// TIA Portal project "ProjektZaliczenie" (V13) (continued)
HMI tags "Default tag table"
   "Player1DataBlock_SelectedSize" : Int, 100 ms
   "Player1DataBlock_Orientation" : Bool, 100 ms
   "Player1DataBlock_ResetAll" : Bool, 100 ms
   "Player1DataBlock_Ready" : Bool, 100 ms
   "Player1DataBlock_SelectedPosition" : Int, 100 ms
   "Player1DataBlock_FieldsTypes" : Array [0..99] of Int, 100 ms
   "Player1DataBlock_Size4Count" : Int, 100 ms
   "Player1DataBlock_Size3Count" : Int, 100 ms
   "Player1DataBlock_Size2Count" : Int, 100 ms
   "Player1DataBlock_Size1Count" : Int, 100 ms
   "Player1DataBlock_ShipsReady" : Bool, 100 ms
   "Tag_ScreenNumber" : UInt, internal
   "MainDataBlock_Turn" : Bool, 100 ms
   "MainDataBlock_GameResult" : Int, 100 ms
   "Player1DataBlock_EnemyBoard{0}" : Int, 100 ms
   "Player1DataBlock_EnemyBoard{1}" : Int, 100 ms
   "Player1DataBlock_EnemyBoard{2}" : Int, 100 ms
   "Player1DataBlock_EnemyBoard{3}" : Int, 100 ms
   "Player1DataBlock_EnemyBoard{4}" : Int, 100 ms
   "Player1DataBlock_EnemyBoard{5}" : Int, 100 ms
   "Player1DataBlock_EnemyBoard{6}" : Int, 100 ms
   "Player1DataBlock_EnemyBoard{7}" : Int, 100 ms
   "Player1DataBlock_EnemyBoard{8}" : Int, 100 ms
   "Player1DataBlock_EnemyBoard{9}" : Int, 100 ms
   "Player1DataBlock_EnemyBoard{10}" : Int, 100 ms
   "Player1DataBlock_EnemyBoard{11}" : Int, 100 ms
   "Player1DataBlock_EnemyBoard{12}" : Int, 100 ms
   "Player1DataBlock_EnemyBoard{13}" : Int, 100 ms
   "Player1DataBlock_EnemyBoard{14}" : Int, 100 ms
   "Player1DataBlock_EnemyBoard{15}" : Int, 100 ms
   "Player1DataBlock_EnemyBoard{16}" : Int, 100 ms
   "Player1DataBlock_EnemyBoard{17}" : Int, 100 ms
   "Player1DataBlock_EnemyBoard{18}" : Int, 100 ms
   "Player1DataBlock_EnemyBoard{19}" : Int, 100 ms
   "Player1DataBlock_EnemyBoard{20}" : Int, 100 ms
   "Player1DataBlock_EnemyBoard{21}" : Int, 100 ms
   "Player1DataBlock_EnemyBoard{22}" : Int, 100 ms
   "Player1DataBlock_EnemyBoard{23}" : Int, 100 ms
   "Player1DataBlock_EnemyBoard{24}" : Int, 100 ms
   "Player1DataBlock_EnemyBoard{25}" : Int, 100 ms
   "Player1DataBlock_EnemyBoard{26}" : Int, 100 ms
   "Player1DataBlock_EnemyBoard{27}" : Int, 100 ms
   "Player1DataBlock_EnemyBoard{28}" : Int, 100 ms
   "Player1DataBlock_EnemyBoard{29}" : Int, 100 ms
   "Player1DataBlock_EnemyBoard{30}" : Int, 100 ms
   "Player1DataBlock_EnemyBoard{31}" : Int, 100 ms
   "Player1DataBlock_EnemyBoard{32}" : Int, 100 ms
   "Player1DataBlock_EnemyBoard{33}" : Int, 100 ms
   "Player1DataBlock_EnemyBoard{34}" : Int, 100 ms
   "Player1DataBlock_EnemyBoard{35}" : Int, 100 ms
   "Player1DataBlock_EnemyBoard{36}" : Int, 100 ms
   "Player1DataBlock_EnemyBoard{37}" : Int, 100 ms
   "Player1DataBlock_EnemyBoard{38}" : Int, 100 ms
   "Player1DataBlock_EnemyBoard{39}" : Int, 100 ms
   "Player1DataBlock_EnemyBoard{40}" : Int, 100 ms
   "Player1DataBlock_EnemyBoard{41}" : Int, 100 ms
   "Player1DataBlock_EnemyBoard{42}" : Int, 100 ms
   "Player1DataBlock_EnemyBoard{43}" : Int, 100 ms
   "Player1DataBlock_EnemyBoard{44}" : Int, 100 ms
   "Player1DataBlock_EnemyBoard{45}" : Int, 100 ms
   "Player1DataBlock_EnemyBoard{46}" : Int, 100 ms
   "Player1DataBlock_EnemyBoard{47}" : Int, 100 ms
   "Player1DataBlock_EnemyBoard{48}" : Int, 100 ms
   "Player1DataBlock_EnemyBoard{49}" : Int, 100 ms
   "Player1DataBlock_EnemyBoard{50}" : Int, 100 ms
   "Player1DataBlock_EnemyBoard{51}" : Int, 100 ms
   "Player1DataBlock_EnemyBoard{52}" : Int, 100 ms
   "Player1DataBlock_EnemyBoard{53}" : Int, 100 ms
   "Player1DataBlock_EnemyBoard{54}" : Int, 100 ms
   "Player1DataBlock_EnemyBoard{55}" : Int, 100 ms
   "Player1DataBlock_EnemyBoard{56}" : Int, 100 ms
   "Player1DataBlock_EnemyBoard{57}" : Int, 100 ms
   "Player1DataBlock_EnemyBoard{58}" : Int, 100 ms
   "Player1DataBlock_EnemyBoard{59}" : Int, 100 ms
   "Player1DataBlock_EnemyBoard{60}" : Int, 100 ms
   "Player1DataBlock_EnemyBoard{61}" : Int, 100 ms
   "Player1DataBlock_EnemyBoard{62}" : Int, 100 ms
   "Player1DataBlock_EnemyBoard{63}" : Int, 100 ms
   "Player1DataBlock_EnemyBoard{64}" : Int, 100 ms
   "Player1DataBlock_EnemyBoard{65}" : Int, 100 ms
   "Player1DataBlock_EnemyBoard{66}" : Int, 100 ms
   "Player1DataBlock_EnemyBoard{67}" : Int, 100 ms
   "Player1DataBlock_EnemyBoard{68}" : Int, 100 ms
   "Player1DataBlock_EnemyBoard{69}" : Int, 100 ms
   "Player1DataBlock_EnemyBoard{70}" : Int, 100 ms
   "Player1DataBlock_EnemyBoard{71}" : Int, 100 ms
   "Player1DataBlock_EnemyBoard{72}" : Int, 100 ms
   "Player1DataBlock_EnemyBoard{73}" : Int, 100 ms
   "Player1DataBlock_EnemyBoard{74}" : Int, 100 ms
   "Player1DataBlock_EnemyBoard{75}" : Int, 100 ms
   "Player1DataBlock_EnemyBoard{76}" : Int, 100 ms
   "Player1DataBlock_EnemyBoard{77}" : Int, 100 ms
   "Player1DataBlock_EnemyBoard{78}" : Int, 100 ms
   "Player1DataBlock_EnemyBoard{79}" : Int, 100 ms
   "Player1DataBlock_EnemyBoard{80}" : Int, 100 ms
   "Player1DataBlock_EnemyBoard{81}" : Int, 100 ms
   "Player1DataBlock_EnemyBoard{82}" : Int, 100 ms
   "Player1DataBlock_EnemyBoard{83}" : Int, 100 ms
   "Player1DataBlock_EnemyBoard{84}" : Int, 100 ms
   "Player1DataBlock_EnemyBoard{85}" : Int, 100 ms
   "Player1DataBlock_EnemyBoard{86}" : Int, 100 ms
   "Player1DataBlock_EnemyBoard{87}" : Int, 100 ms
   "Player1DataBlock_EnemyBoard{88}" : Int, 100 ms
   "Player1DataBlock_EnemyBoard{89}" : Int, 100 ms
   "Player1DataBlock_EnemyBoard{90}" : Int, 100 ms
   "Player1DataBlock_EnemyBoard{91}" : Int, 100 ms
   "Player1DataBlock_EnemyBoard{92}" : Int, 100 ms
   "Player1DataBlock_EnemyBoard{93}" : Int, 100 ms
   "Player1DataBlock_EnemyBoard{94}" : Int, 100 ms
   "Player1DataBlock_EnemyBoard{95}" : Int, 100 ms
   "Player1DataBlock_EnemyBoard{96}" : Int, 100 ms
   "Player1DataBlock_EnemyBoard{97}" : Int, 100 ms
   "Player1DataBlock_EnemyBoard{98}" : Int, 100 ms
   "Player1DataBlock_EnemyBoard{99}" : Int, 100 ms
   "Player1DataBlock_ReadyForNewGame" : Bool, 100 ms
   "Player1DataBlock_GraphicsTypes" : Array [0..99] of Int, 100 ms
   "MainDataBlock_Player2Won" : Bool, 1 s
   "MainDataBlock_Player1Won" : Bool, 1 s

text list "gameResults": 0 ''; 1 ''; 2 ''

graphic list "Player": 2 'blue'; 0 'blue'; 1 'statek1_1'; 3 'statek1_red'; 20 'statek2_2'; 31 'statek31'; 32 'statek32'; 33 'statek33'; 41 'statek41'; 42 'statek42'; 43 'statek43'; 44 'statek44'; 101 'statek101'; 201 'statek101_1'; 202 'statek202'; 301 'statek301'; 302 'statek302'; 303 'statek303'; 401 'statek401'; 402 'statek402'; 403 'statek403'; 404 'statek404'; 333 'hit'; 444 'boom_1'

graphic list "Enemy": 0 'enemy_un'; 3 'boom_1'; 2 'hit'

screen "Stage2" 800x480, template "Template_1"
   Button "Button_1" at 39,131 size 32x32
   GraphicView "Graphic view_3" at 0,0 size 800x479
   GraphicView "Graphic view_2" at 410,97 size 376x366
   GraphicView "Graphic view_1" at 2,95 size 378x366
   Button "Button_101" at 445,131 size 32x32
   Button "Button_102" at 479,131 size 32x32
   Button "Button_103" at 513,131 size 32x32
   Button "Button_104" at 547,131 size 32x32
   Button "Button_105" at 581,131 size 32x32
   Button "Button_106" at 615,131 size 32x32
   Button "Button_107" at 649,131 size 32x32
   Button "Button_108" at 683,131 size 32x32
   Button "Button_109" at 717,131 size 32x32
   Button "Button_110" at 751,131 size 32x32
   Button "Button_111" at 445,164 size 32x32
   Button "Button_112" at 479,164 size 32x32
   Button "Button_113" at 513,164 size 32x32
   Button "Button_114" at 547,164 size 32x32
   Button "Button_115" at 581,164 size 32x32
   Button "Button_116" at 615,164 size 32x32
   Button "Button_117" at 649,164 size 32x32
   Button "Button_118" at 683,164 size 32x32
   Button "Button_119" at 717,164 size 32x32
   Button "Button_120" at 751,164 size 32x32
   Button "Button_121" at 445,197 size 32x32
   Button "Button_122" at 479,197 size 32x32
   Button "Button_123" at 513,197 size 32x32
   Button "Button_124" at 547,197 size 32x32
   Button "Button_125" at 581,197 size 32x32
   Button "Button_126" at 615,197 size 32x32
   Button "Button_127" at 649,197 size 32x32
   Button "Button_128" at 683,197 size 32x32
   Button "Button_129" at 717,197 size 32x32
   Button "Button_130" at 751,197 size 32x32
   Button "Button_131" at 445,230 size 32x32
   Button "Button_132" at 479,230 size 32x32
   Button "Button_133" at 513,230 size 32x32
   Button "Button_134" at 547,230 size 32x32
   Button "Button_135" at 581,230 size 32x32
   Button "Button_136" at 615,230 size 32x32
   Button "Button_137" at 649,230 size 32x32
   Button "Button_138" at 683,230 size 32x32
   Button "Button_139" at 717,230 size 32x32
   Button "Button_140" at 751,230 size 32x32
   Button "Button_141" at 445,263 size 32x32
   Button "Button_142" at 479,263 size 32x32
   Button "Button_143" at 513,263 size 32x32
   Button "Button_144" at 547,263 size 32x32
   Button "Button_145" at 581,263 size 32x32
   Button "Button_146" at 615,263 size 32x32
   Button "Button_147" at 649,263 size 32x32
   Button "Button_148" at 683,263 size 32x32
   Button "Button_149" at 717,263 size 32x32
   Button "Button_150" at 751,263 size 32x32
   Button "Button_151" at 445,296 size 32x32
   Button "Button_152" at 479,296 size 32x32
   Button "Button_153" at 513,296 size 32x32
   Button "Button_154" at 547,296 size 32x32
   Button "Button_155" at 581,296 size 32x32
   Button "Button_156" at 615,296 size 32x32
   Button "Button_157" at 649,296 size 32x32
   Button "Button_158" at 683,296 size 32x32
   Button "Button_159" at 717,296 size 32x32
   Button "Button_160" at 751,296 size 32x32
   Button "Button_161" at 445,329 size 32x32
   Button "Button_162" at 479,329 size 32x32
   Button "Button_163" at 513,329 size 32x32
   Button "Button_164" at 547,329 size 32x32
   Button "Button_165" at 581,329 size 32x32
   Button "Button_166" at 615,329 size 32x32
   Button "Button_167" at 649,329 size 32x32
   Button "Button_168" at 683,329 size 32x32
   Button "Button_169" at 717,329 size 32x32
   Button "Button_170" at 751,329 size 32x32
   Button "Button_171" at 445,362 size 32x32
   Button "Button_172" at 479,362 size 32x32
   Button "Button_173" at 513,362 size 32x32
   Button "Button_174" at 547,362 size 32x32
   Button "Button_175" at 581,362 size 32x32
   Button "Button_176" at 615,362 size 32x32
   Button "Button_177" at 649,362 size 32x32
   Button "Button_178" at 683,362 size 32x32
   Button "Button_179" at 717,362 size 32x32
   Button "Button_180" at 751,362 size 32x32
   Button "Button_181" at 445,395 size 32x32
   Button "Button_182" at 479,395 size 32x32
   Button "Button_183" at 513,395 size 32x32
   Button "Button_184" at 547,395 size 32x32
   Button "Button_185" at 581,395 size 32x32
   Button "Button_186" at 615,395 size 32x32
   Button "Button_187" at 649,395 size 32x32
   Button "Button_188" at 683,395 size 32x32
   Button "Button_189" at 717,395 size 32x32
   Button "Button_190" at 751,395 size 32x32
   Button "Button_191" at 445,428 size 32x32
   Button "Button_192" at 479,428 size 32x32
   Button "Button_193" at 513,428 size 32x32
   Button "Button_194" at 547,428 size 32x32
   Button "Button_195" at 581,428 size 32x32
   Button "Button_196" at 615,428 size 32x32
   Button "Button_197" at 649,428 size 32x32
   Button "Button_198" at 683,428 size 32x32
   Button "Button_199" at 717,428 size 32x32
   Button "Button_200" at 751,428 size 32x32
   TextField "Text field_41" at 144,72 size 100x23
   TextField "Text field_42" at 556,72 size 140x23
   TextField "Text field_43" at 372,11 size 76x23
   Button "Button_201" at 721,8 size 33x20
   Button "Button_202" at 721,31 size 33x20
   Button "Button_203" at 721,56 size 33x20
   Button "Button_2" at 73,130 size 32x32
   Button "Button_3" at 107,130 size 32x32
   Button "Button_4" at 141,130 size 32x32
   Button "Button_5" at 175,130 size 32x32
   Button "Button_6" at 209,130 size 32x32
   Button "Button_7" at 243,130 size 32x32
   Button "Button_8" at 277,130 size 32x32
   Button "Button_9" at 311,130 size 32x32
   Button "Button_10" at 345,130 size 32x32
   Button "Button_11" at 39,163 size 32x32
   Button "Button_12" at 73,163 size 32x32
   Button "Button_13" at 107,163 size 32x32
   Button "Button_14" at 141,163 size 32x32
   Button "Button_15" at 175,163 size 32x32
   Button "Button_16" at 209,163 size 32x32
   Button "Button_17" at 243,163 size 32x32
   Button "Button_18" at 277,163 size 32x32
   Button "Button_19" at 311,163 size 32x32
   Button "Button_20" at 345,163 size 32x32
   Button "Button_21" at 39,196 size 32x32
   Button "Button_22" at 73,196 size 32x32
   Button "Button_23" at 107,196 size 32x32
   Button "Button_24" at 141,196 size 32x32
   Button "Button_25" at 175,196 size 32x32
   Button "Button_26" at 209,196 size 32x32
   Button "Button_27" at 243,196 size 32x32
   Button "Button_28" at 277,196 size 32x32
   Button "Button_29" at 311,196 size 32x32
   Button "Button_30" at 345,196 size 32x32
   Button "Button_31" at 39,229 size 32x32
   Button "Button_32" at 73,229 size 32x32
   Button "Button_33" at 107,229 size 32x32
   Button "Button_34" at 141,229 size 32x32
   Button "Button_35" at 175,229 size 32x32
   Button "Button_36" at 209,229 size 32x32
   Button "Button_37" at 243,229 size 32x32
   Button "Button_38" at 277,229 size 32x32
   Button "Button_39" at 311,229 size 32x32
   Button "Button_40" at 345,229 size 32x32
   Button "Button_41" at 39,262 size 32x32
   Button "Button_42" at 73,262 size 32x32
   Button "Button_43" at 107,262 size 32x32
   Button "Button_44" at 141,262 size 32x32
   Button "Button_45" at 175,262 size 32x32
   Button "Button_46" at 209,262 size 32x32
   Button "Button_47" at 243,262 size 32x32
   Button "Button_48" at 277,262 size 32x32
   Button "Button_49" at 311,262 size 32x32
   Button "Button_50" at 345,262 size 32x32
   Button "Button_51" at 39,295 size 32x32
   Button "Button_52" at 73,295 size 32x32
   Button "Button_53" at 107,295 size 32x32
   Button "Button_54" at 141,295 size 32x32
   Button "Button_55" at 175,295 size 32x32
   Button "Button_56" at 209,295 size 32x32
   Button "Button_57" at 243,295 size 32x32
   Button "Button_58" at 277,295 size 32x32
   Button "Button_59" at 311,295 size 32x32
   Button "Button_60" at 345,295 size 32x32
   Button "Button_61" at 39,328 size 32x32
   Button "Button_62" at 73,328 size 32x32
   Button "Button_63" at 107,328 size 32x32
   Button "Button_64" at 141,328 size 32x32
   Button "Button_65" at 175,328 size 32x32
   Button "Button_66" at 209,328 size 32x32
   Button "Button_67" at 243,328 size 32x32
   Button "Button_68" at 277,328 size 32x32
   Button "Button_69" at 311,328 size 32x32
   Button "Button_70" at 345,328 size 32x32
   Button "Button_71" at 39,361 size 32x32
   Button "Button_72" at 73,361 size 32x32
   Button "Button_73" at 107,361 size 32x32
   Button "Button_74" at 141,361 size 32x32
   Button "Button_75" at 175,361 size 32x32
   Button "Button_76" at 209,361 size 32x32
   Button "Button_77" at 243,361 size 32x32
   Button "Button_78" at 277,361 size 32x32
   Button "Button_79" at 311,361 size 32x32
   Button "Button_81" at 39,394 size 32x32
   Button "Button_82" at 73,394 size 32x32
   Button "Button_83" at 107,394 size 32x32
   Button "Button_84" at 141,394 size 32x32
   Button "Button_85" at 175,394 size 32x32
   Button "Button_86" at 209,394 size 32x32
   Button "Button_87" at 243,394 size 32x32
   Button "Button_88" at 277,394 size 32x32
   Button "Button_89" at 311,394 size 32x32
   Button "Button_90" at 345,394 size 32x32
   Button "Button_91" at 39,427 size 32x32
   Button "Button_92" at 73,427 size 32x32
   Button "Button_93" at 107,427 size 32x32
   Button "Button_94" at 141,427 size 32x32
   Button "Button_95" at 175,427 size 32x32
   Button "Button_96" at 209,427 size 32x32
   Button "Button_97" at 243,427 size 32x32
   Button "Button_98" at 277,427 size 32x32
   Button "Button_99" at 311,427 size 32x32
   Button "Button_100" at 345,427 size 32x32
   Button "Button_80" at 345,361 size 32x32

screen "Stage1" 800x480
   Button "Button_1" at 39,131 size 32x32
   GraphicView "Graphic view_1" at 0,0 size 799x479
   GraphicView "Graphic view_2" at 0,96 size 381x363
   Button "Button_2" at 73,130 size 32x32
   Button "Button_3" at 107,130 size 32x32
   Button "Button_4" at 141,130 size 32x32
   Button "Button_5" at 175,130 size 32x32
   Button "Button_6" at 209,130 size 32x32
   Button "Button_7" at 243,130 size 32x32
   Button "Button_8" at 277,130 size 32x32
   Button "Button_9" at 311,130 size 32x32
   Button "Button_10" at 345,130 size 32x32
   Button "Button_11" at 39,163 size 32x32
   Button "Button_12" at 73,163 size 32x32
   Button "Button_13" at 107,163 size 32x32
   Button "Button_14" at 141,163 size 32x32
   Button "Button_15" at 175,163 size 32x32
   Button "Button_16" at 209,163 size 32x32
   Button "Button_17" at 243,163 size 32x32
   Button "Button_18" at 277,163 size 32x32
   Button "Button_19" at 311,163 size 32x32
   Button "Button_20" at 345,163 size 32x32
   Button "Button_21" at 39,196 size 32x32
   Button "Button_22" at 73,196 size 32x32
   Button "Button_23" at 107,196 size 32x32
   Button "Button_24" at 141,196 size 32x32
   Button "Button_25" at 175,196 size 32x32
   Button "Button_26" at 209,196 size 32x32
   Button "Button_27" at 243,196 size 32x32
   Button "Button_28" at 277,196 size 32x32
   Button "Button_29" at 311,196 size 32x32
   Button "Button_30" at 345,196 size 32x32
   Button "Button_31" at 39,229 size 32x32
   Button "Button_32" at 73,229 size 32x32
   Button "Button_33" at 107,229 size 32x32
   Button "Button_34" at 141,229 size 32x32
   Button "Button_35" at 175,229 size 32x32
   Button "Button_36" at 209,229 size 32x32
   Button "Button_37" at 243,229 size 32x32
   Button "Button_38" at 277,229 size 32x32
   Button "Button_39" at 311,229 size 32x32
   Button "Button_40" at 345,229 size 32x32
   Button "Button_41" at 39,262 size 32x32
   Button "Button_42" at 73,262 size 32x32
   Button "Button_43" at 107,262 size 32x32
   Button "Button_44" at 141,262 size 32x32
   Button "Button_45" at 175,262 size 32x32
   Button "Button_46" at 209,262 size 32x32
   Button "Button_47" at 243,262 size 32x32
   Button "Button_48" at 277,262 size 32x32
   Button "Button_49" at 311,262 size 32x32
   Button "Button_50" at 345,262 size 32x32
   Button "Button_51" at 39,295 size 32x32
   Button "Button_52" at 73,295 size 32x32
   Button "Button_53" at 107,295 size 32x32
   Button "Button_54" at 141,295 size 32x32
   Button "Button_55" at 175,295 size 32x32
   Button "Button_56" at 209,295 size 32x32
   Button "Button_57" at 243,295 size 32x32
   Button "Button_58" at 277,295 size 32x32
   Button "Button_59" at 311,295 size 32x32
   Button "Button_60" at 345,295 size 32x32
   Button "Button_61" at 39,328 size 32x32
   Button "Button_62" at 73,328 size 32x32
   Button "Button_63" at 107,328 size 32x32
   Button "Button_64" at 141,328 size 32x32
   Button "Button_65" at 175,328 size 32x32
   Button "Button_66" at 209,328 size 32x32
   Button "Button_67" at 243,328 size 32x32
   Button "Button_68" at 277,328 size 32x32
   Button "Button_69" at 311,328 size 32x32
   Button "Button_70" at 345,328 size 32x32
   Button "Button_71" at 39,361 size 32x32
   Button "Button_72" at 73,361 size 32x32
   Button "Button_73" at 107,361 size 32x32
   Button "Button_74" at 141,361 size 32x32
   Button "Button_75" at 175,361 size 32x32
   Button "Button_76" at 209,361 size 32x32
   Button "Button_77" at 243,361 size 32x32
   Button "Button_78" at 277,361 size 32x32
   Button "Button_79" at 311,361 size 32x32
   Button "Button_81" at 39,394 size 32x32
   Button "Button_82" at 73,394 size 32x32
   Button "Button_83" at 107,394 size 32x32
   Button "Button_84" at 141,394 size 32x32
   Button "Button_85" at 175,394 size 32x32
   Button "Button_86" at 209,394 size 32x32
   Button "Button_87" at 243,394 size 32x32
   Button "Button_88" at 277,394 size 32x32
   Button "Button_89" at 311,394 size 32x32
   Button "Button_90" at 345,394 size 32x32
   Button "Button_91" at 39,427 size 32x32
   Button "Button_92" at 73,427 size 32x32
   Button "Button_93" at 107,427 size 32x32
   Button "Button_94" at 141,427 size 32x32
   Button "Button_95" at 175,427 size 32x32
   Button "Button_96" at 209,427 size 32x32
   Button "Button_97" at 243,427 size 32x32
   Button "Button_98" at 277,427 size 32x32
   Button "Button_99" at 311,427 size 32x32
   Button "Button_100" at 345,427 size 32x32
   Button "Button_80" at 345,361 size 32x32
   Switch "Switch_1" at 643,281 size 131x41
   Button "Button_101" at 417,142 size 134x32
   Button "Button_102" at 417,181 size 103x37
   Button "Button_103" at 417,233 size 66x32
   Button "Button_104" at 417,281 size 32x32
   Button "Button_105" at 611,135 size 164x46
   Switch "Switch_2" at 597,403 size 178x44
   TextField "Text field_21" at 296,36 size 232x23
   Button "Button_106" at 742,16 size 33x20
   Button "Button_107" at 742,36 size 33x20
   Button "Button_108" at 741,59 size 33x20

screen "Stage3" 800x480
   GraphicView "Graphic view_1" at 0,0 size 799x479
   Button "Button_1" at 265,294 size 282x65
   Button "Button_106" at 643,36 size 33x20
   Button "Button_107" at 682,36 size 33x20
   Button "Button_108" at 721,36 size 33x20
   Button "Button_2" at 253,139 size 305x32
*)

(* ===== HMI "HMI_RT_3" =====
connection "HMI_Connection_3": ETHERNET, SMART_S7_1200_OMS

HMI tags "Default tag table"
   "Player2DataBlock_GraphicsTypes" : Array [0..99] of Int, 100 ms
   "Player2DataBlock_SelectedPosition" : Int, 100 ms
   "Player2DataBlock_FieldsTypes" : Array [0..99] of Int, 100 ms
   "Player2DataBlock_Orientation" : Bool, 100 ms
   "Player2DataBlock_PlayerReady" : Bool, 100 ms
   "Player2DataBlock_ResetAll" : Bool, 100 ms
   "Player2DataBlock_SelectedSize" : Int, 100 ms
   "Player2DataBlock_ShipsReady" : Bool, 100 ms
   "Player2DataBlock_Size1Count" : Int, 100 ms
   "Player2DataBlock_Size2Count" : Int, 100 ms
   "Player2DataBlock_Size3Count" : Int, 100 ms
   "Player2DataBlock_Size4Count" : Int, 100 ms
   "MainDataBlock_Turn" : Bool, 100 ms
   "MainDataBlock_GameResult" : Int, 100 ms
   "Player2DataBlock_EnemyBoard{0}" : Int, 100 ms
   "Player2DataBlock_EnemyBoard{1}" : Int, 100 ms
   "Player2DataBlock_EnemyBoard{2}" : Int, 100 ms
   "Player2DataBlock_EnemyBoard{3}" : Int, 100 ms
   "Player2DataBlock_EnemyBoard{4}" : Int, 100 ms
   "Player2DataBlock_EnemyBoard{5}" : Int, 100 ms
   "Player2DataBlock_EnemyBoard{6}" : Int, 100 ms
   "Player2DataBlock_EnemyBoard{7}" : Int, 100 ms
   "Player2DataBlock_EnemyBoard{8}" : Int, 100 ms
   "Player2DataBlock_EnemyBoard{9}" : Int, 100 ms
   "Player2DataBlock_EnemyBoard{10}" : Int, 100 ms
   "Player2DataBlock_EnemyBoard{11}" : Int, 100 ms
   "Player2DataBlock_EnemyBoard{12}" : Int, 100 ms
   "Player2DataBlock_EnemyBoard{13}" : Int, 100 ms
   "Player2DataBlock_EnemyBoard{14}" : Int, 100 ms
   "Player2DataBlock_EnemyBoard{15}" : Int, 100 ms
   "Player2DataBlock_EnemyBoard{16}" : Int, 100 ms
   "Player2DataBlock_EnemyBoard{17}" : Int, 100 ms
   "Player2DataBlock_EnemyBoard{18}" : Int, 100 ms
   "Player2DataBlock_EnemyBoard{19}" : Int, 100 ms
   "Player2DataBlock_EnemyBoard{20}" : Int, 100 ms
   "Player2DataBlock_EnemyBoard{21}" : Int, 100 ms
   "Player2DataBlock_EnemyBoard{22}" : Int, 100 ms
   "Player2DataBlock_EnemyBoard{23}" : Int, 100 ms
   "Player2DataBlock_EnemyBoard{24}" : Int, 100 ms
   "Player2DataBlock_EnemyBoard{25}" : Int, 100 ms
   "Player2DataBlock_EnemyBoard{26}" : Int, 100 ms
   "Player2DataBlock_EnemyBoard{27}" : Int, 100 ms
   "Player2DataBlock_EnemyBoard{28}" : Int, 100 ms
   "Player2DataBlock_EnemyBoard{29}" : Int, 100 ms
   "Player2DataBlock_EnemyBoard{30}" : Int, 100 ms
   "Player2DataBlock_EnemyBoard{31}" : Int, 100 ms
   "Player2DataBlock_EnemyBoard{32}" : Int, 100 ms
   "Player2DataBlock_EnemyBoard{33}" : Int, 100 ms
   "Player2DataBlock_EnemyBoard{34}" : Int, 100 ms
   "Player2DataBlock_EnemyBoard{35}" : Int, 100 ms
   "Player2DataBlock_EnemyBoard{36}" : Int, 100 ms
   "Player2DataBlock_EnemyBoard{37}" : Int, 100 ms
   "Player2DataBlock_EnemyBoard{38}" : Int, 100 ms
   "Player2DataBlock_EnemyBoard{39}" : Int, 100 ms
   "Player2DataBlock_EnemyBoard{40}" : Int, 100 ms
   "Player2DataBlock_EnemyBoard{41}" : Int, 100 ms
   "Player2DataBlock_EnemyBoard{42}" : Int, 100 ms
   "Player2DataBlock_EnemyBoard{43}" : Int, 100 ms
   "Player2DataBlock_EnemyBoard{44}" : Int, 100 ms
   "Player2DataBlock_EnemyBoard{45}" : Int, 100 ms
   "Player2DataBlock_EnemyBoard{46}" : Int, 100 ms
   "Player2DataBlock_EnemyBoard{47}" : Int, 100 ms
   "Player2DataBlock_EnemyBoard{48}" : Int, 100 ms
   "Player2DataBlock_EnemyBoard{49}" : Int, 100 ms
   "Player2DataBlock_EnemyBoard{50}" : Int, 100 ms
   "Player2DataBlock_EnemyBoard{51}" : Int, 100 ms
   "Player2DataBlock_EnemyBoard{52}" : Int, 100 ms
   "Player2DataBlock_EnemyBoard{53}" : Int, 100 ms
   "Player2DataBlock_EnemyBoard{54}" : Int, 100 ms
   "Player2DataBlock_EnemyBoard{55}" : Int, 100 ms
   "Player2DataBlock_EnemyBoard{56}" : Int, 100 ms
   "Player2DataBlock_EnemyBoard{57}" : Int, 100 ms
   "Player2DataBlock_EnemyBoard{58}" : Int, 100 ms
   "Player2DataBlock_EnemyBoard{59}" : Int, 100 ms
   "Player2DataBlock_EnemyBoard{60}" : Int, 100 ms
   "Player2DataBlock_EnemyBoard{61}" : Int, 100 ms
   "Player2DataBlock_EnemyBoard{62}" : Int, 100 ms
   "Player2DataBlock_EnemyBoard{63}" : Int, 100 ms
   "Player2DataBlock_EnemyBoard{64}" : Int, 100 ms
   "Player2DataBlock_EnemyBoard{65}" : Int, 100 ms
   "Player2DataBlock_EnemyBoard{66}" : Int, 100 ms
   "Player2DataBlock_EnemyBoard{67}" : Int, 100 ms
   "Player2DataBlock_EnemyBoard{68}" : Int, 100 ms
   "Player2DataBlock_EnemyBoard{69}" : Int, 100 ms
   "Player2DataBlock_EnemyBoard{70}" : Int, 100 ms
   "Player2DataBlock_EnemyBoard{71}" : Int, 100 ms
   "Player2DataBlock_EnemyBoard{72}" : Int, 100 ms
   "Player2DataBlock_EnemyBoard{73}" : Int, 100 ms
   "Player2DataBlock_EnemyBoard{74}" : Int, 100 ms
   "Player2DataBlock_EnemyBoard{75}" : Int, 100 ms
   "Player2DataBlock_EnemyBoard{76}" : Int, 100 ms
   "Player2DataBlock_EnemyBoard{77}" : Int, 100 ms
   "Player2DataBlock_EnemyBoard{78}" : Int, 100 ms
   "Player2DataBlock_EnemyBoard{79}" : Int, 100 ms
   "Player2DataBlock_EnemyBoard{80}" : Int, 100 ms
   "Player2DataBlock_EnemyBoard{81}" : Int, 100 ms
   "Player2DataBlock_EnemyBoard{82}" : Int, 100 ms
   "Player2DataBlock_EnemyBoard{83}" : Int, 100 ms
   "Player2DataBlock_EnemyBoard{84}" : Int, 100 ms
   "Player2DataBlock_EnemyBoard{85}" : Int, 100 ms
   "Player2DataBlock_EnemyBoard{86}" : Int, 100 ms
   "Player2DataBlock_EnemyBoard{87}" : Int, 100 ms
   "Player2DataBlock_EnemyBoard{88}" : Int, 100 ms
   "Player2DataBlock_EnemyBoard{89}" : Int, 100 ms
   "Player2DataBlock_EnemyBoard{90}" : Int, 100 ms
   "Player2DataBlock_EnemyBoard{91}" : Int, 100 ms
   "Player2DataBlock_EnemyBoard{92}" : Int, 100 ms
   "Player2DataBlock_EnemyBoard{93}" : Int, 100 ms
   "Player2DataBlock_EnemyBoard{94}" : Int, 100 ms
   "Player2DataBlock_EnemyBoard{95}" : Int, 100 ms
   "Player2DataBlock_EnemyBoard{96}" : Int, 100 ms
   "Player2DataBlock_EnemyBoard{97}" : Int, 100 ms
   "Player2DataBlock_EnemyBoard{98}" : Int, 100 ms
   "Player2DataBlock_EnemyBoard{99}" : Int, 100 ms
   "Player2DataBlock_ReadyForNewGame" : Bool, 100 ms
   "MainDataBlock_Player2Won" : Bool, 1 s
   "MainDataBlock_Player1Won" : Bool, 1 s

text list "gameResults": 0 ''; 1 ''; 2 ''

graphic list "Graphic_list_2": 2 'blue'; 0 'blue'; 1 'statek1_1'; 3 'statek1_red'; 20 'statek2_2'; 31 'statek31'; 32 'statek32'; 33 'statek33'; 41 'statek41'; 42 'statek42'; 43 'statek43'; 44 'statek44'; 101 'statek101'; 201 'statek101_1'; 202 'statek202'; 301 'statek301'; 302 'statek302'; 303 'statek303'; 401 'statek401'; 402 'statek402'; 403 'statek403'; 404 'statek404'; 333 'hit'; 444 'boom_1'

graphic list "Enemy": 0 'enemy_un'; 3 'boom_1'; 2 'hit'

screen "Stage1" 800x480
   GraphicView "Graphic view_1" at 0,0 size 800x480
   GraphicView "Graphic view_2" at 0,95 size 382x366
   Button "Button_1" at 39,130 size 32x32
   Button "Button_2" at 73,130 size 32x32
   Button "Button_3" at 107,130 size 32x32
   Button "Button_4" at 141,130 size 32x32
   Button "Button_5" at 175,130 size 32x32
   Button "Button_6" at 209,130 size 32x32
   Button "Button_7" at 243,130 size 32x32
   Button "Button_8" at 277,130 size 32x32
   Button "Button_9" at 311,130 size 32x32
   Button "Button_10" at 345,130 size 32x32
   Button "Button_11" at 39,163 size 32x32
   Button "Button_12" at 73,163 size 32x32
   Button "Button_13" at 107,163 size 32x32
   Button "Button_14" at 141,163 size 32x32
   Button "Button_15" at 175,163 size 32x32
   Button "Button_16" at 209,163 size 32x32
   Button "Button_17" at 243,163 size 32x32
   Button "Button_18" at 277,163 size 32x32
   Button "Button_19" at 311,163 size 32x32
   Button "Button_20" at 345,163 size 32x32
   Button "Button_21" at 39,196 size 32x32
   Button "Button_22" at 73,196 size 32x32
   Button "Button_23" at 107,196 size 32x32
   Button "Button_24" at 141,196 size 32x32
   Button "Button_25" at 175,196 size 32x32
   Button "Button_26" at 209,196 size 32x32
   Button "Button_27" at 243,196 size 32x32
   Button "Button_28" at 277,196 size 32x32
   Button "Button_29" at 311,196 size 32x32
   Button "Button_30" at 345,196 size 32x32
   Button "Button_31" at 39,229 size 32x32
   Button "Button_32" at 73,229 size 32x32
   Button "Button_33" at 107,229 size 32x32
   Button "Button_34" at 141,229 size 32x32
   Button "Button_35" at 175,229 size 32x32
   Button "Button_36" at 209,229 size 32x32
   Button "Button_37" at 243,229 size 32x32
   Button "Button_38" at 277,229 size 32x32
   Button "Button_39" at 311,229 size 32x32
   Button "Button_40" at 345,229 size 32x32
   Button "Button_41" at 39,262 size 32x32
   Button "Button_42" at 73,262 size 32x32
   Button "Button_43" at 107,262 size 32x32
   Button "Button_44" at 141,262 size 32x32
   Button "Button_45" at 175,262 size 32x32
   Button "Button_46" at 209,262 size 32x32
   Button "Button_47" at 243,262 size 32x32
   Button "Button_48" at 277,262 size 32x32
   Button "Button_49" at 311,262 size 32x32
   Button "Button_50" at 345,262 size 32x32
   Button "Button_51" at 39,295 size 32x32
   Button "Button_52" at 73,295 size 32x32
   Button "Button_53" at 107,295 size 32x32
   Button "Button_54" at 141,295 size 32x32
   Button "Button_55" at 175,295 size 32x32
   Button "Button_56" at 209,295 size 32x32
   Button "Button_57" at 243,295 size 32x32
   Button "Button_58" at 277,295 size 32x32
   Button "Button_59" at 311,295 size 32x32
   Button "Button_60" at 345,295 size 32x32
   Button "Button_61" at 39,328 size 32x32
   Button "Button_62" at 73,328 size 32x32
   Button "Button_63" at 107,328 size 32x32
   Button "Button_64" at 141,328 size 32x32
   Button "Button_65" at 175,328 size 32x32
   Button "Button_66" at 209,328 size 32x32
   Button "Button_67" at 243,328 size 32x32
   Button "Button_68" at 277,328 size 32x32
   Button "Button_69" at 311,328 size 32x32
   Button "Button_70" at 345,328 size 32x32
   Button "Button_71" at 39,361 size 32x32
   Button "Button_72" at 73,361 size 32x32
   Button "Button_73" at 107,361 size 32x32
   Button "Button_74" at 141,361 size 32x32
   Button "Button_75" at 175,361 size 32x32
   Button "Button_76" at 209,361 size 32x32
   Button "Button_77" at 243,361 size 32x32
   Button "Button_78" at 277,361 size 32x32
   Button "Button_79" at 311,361 size 32x32
   Button "Button_80" at 345,361 size 32x32
   Button "Button_81" at 39,394 size 32x32
   Button "Button_82" at 73,394 size 32x32
   Button "Button_83" at 107,394 size 32x32
   Button "Button_84" at 141,394 size 32x32
   Button "Button_85" at 175,394 size 32x32
   Button "Button_86" at 209,394 size 32x32
   Button "Button_87" at 243,394 size 32x32
   Button "Button_88" at 277,394 size 32x32
   Button "Button_89" at 311,394 size 32x32
   Button "Button_90" at 345,394 size 32x32
   Button "Button_91" at 39,427 size 32x32
   Button "Button_92" at 73,427 size 32x32
   Button "Button_93" at 107,427 size 32x32
   Button "Button_94" at 141,427 size 32x32
   Button "Button_95" at 175,427 size 32x32
   Button "Button_96" at 209,427 size 32x32
   Button "Button_97" at 243,427 size 32x32
   Button "Button_98" at 277,427 size 32x32
   Button "Button_99" at 311,427 size 32x32
   Button "Button_100" at 345,427 size 32x32
   TextField "Text field_21" at 296,36 size 232x23
   Switch "Switch_1" at 640,284 size 131x41
   Button "Button_101" at 416,144 size 134x32
   Button "Button_102" at 416,186 size 100x32
   Button "Button_103" at 416,229 size 67x34
   Button "Button_104" at 422,284 size 32x32
   Button "Button_105" at 614,134 size 164x46
   Switch "Switch_2" at 602,403 size 178x44
   Button "Button_106" at 747,18 size 33x20
   Button "Button_107" at 745,36 size 33x20
   Button "Button_108" at 747,56 size 33x20

screen "Stage3" 800x480
   GraphicView "Graphic view_1" at 0,0 size 799x479
   Button "Button_1" at 265,294 size 282x65
   Button "Button_106" at 643,36 size 33x20
   Button "Button_107" at 682,36 size 33x20
   Button "Button_108" at 721,36 size 33x20
   Button "Button_2" at 253,139 size 305x32

screen "Stage2" 800x480
   GraphicView "Graphic view_3" at 0,0 size 799x479
   GraphicView "Graphic view_1" at 1,95 size 378x366
   TextField "Text field_41" at 145,70 size 100x23
   TextField "Text field_42" at 562,70 size 140x23
   TextField "Text field_43" at 371,12 size 76x23
   Button "Button_201" at 720,14 size 33x20
   Button "Button_202" at 720,37 size 33x20
   Button "Button_203" at 720,58 size 33x20
   Button "Button_1" at 39,130 size 32x32
   Button "Button_2" at 73,130 size 32x32
   Button "Button_3" at 107,130 size 32x32
   Button "Button_4" at 141,130 size 32x32
   Button "Button_5" at 175,130 size 32x32
   Button "Button_6" at 209,130 size 32x32
   Button "Button_7" at 243,130 size 32x32
   Button "Button_8" at 277,130 size 32x32
   Button "Button_9" at 311,130 size 32x32
   Button "Button_10" at 345,130 size 32x32
   Button "Button_11" at 39,163 size 32x32
   Button "Button_12" at 73,163 size 32x32
   Button "Button_13" at 107,163 size 32x32
   Button "Button_14" at 141,163 size 32x32
   Button "Button_15" at 175,163 size 32x32
   Button "Button_16" at 209,163 size 32x32
   Button "Button_17" at 243,163 size 32x32
   Button "Button_18" at 277,163 size 32x32
   Button "Button_19" at 311,163 size 32x32
   Button "Button_20" at 345,163 size 32x32
   Button "Button_21" at 39,196 size 32x32
   Button "Button_22" at 73,196 size 32x32
   Button "Button_23" at 107,196 size 32x32
   Button "Button_24" at 141,196 size 32x32
   Button "Button_25" at 175,196 size 32x32
   Button "Button_26" at 209,196 size 32x32
   Button "Button_27" at 243,196 size 32x32
   Button "Button_28" at 277,196 size 32x32
   Button "Button_29" at 311,196 size 32x32
   Button "Button_30" at 345,196 size 32x32
   Button "Button_31" at 39,229 size 32x32
   Button "Button_32" at 73,229 size 32x32
   Button "Button_33" at 107,229 size 32x32
   Button "Button_34" at 141,229 size 32x32
   Button "Button_35" at 175,229 size 32x32
   Button "Button_36" at 209,229 size 32x32
   Button "Button_37" at 243,229 size 32x32
   Button "Button_38" at 277,229 size 32x32
   Button "Button_39" at 311,229 size 32x32
   Button "Button_40" at 345,229 size 32x32
   Button "Button_41" at 39,262 size 32x32
   Button "Button_42" at 73,262 size 32x32
   Button "Button_43" at 107,262 size 32x32
   Button "Button_44" at 141,262 size 32x32
   Button "Button_45" at 175,262 size 32x32
   Button "Button_46" at 209,262 size 32x32
   Button "Button_47" at 243,262 size 32x32
   Button "Button_48" at 277,262 size 32x32
   Button "Button_49" at 311,262 size 32x32
   Button "Button_50" at 345,262 size 32x32
   Button "Button_51" at 39,295 size 32x32
   Button "Button_52" at 73,295 size 32x32
   Button "Button_53" at 107,295 size 32x32
   Button "Button_54" at 141,295 size 32x32
   Button "Button_55" at 175,295 size 32x32
   Button "Button_56" at 209,295 size 32x32
   Button "Button_57" at 243,295 size 32x32
   Button "Button_58" at 277,295 size 32x32
   Button "Button_59" at 311,295 size 32x32
   Button "Button_60" at 345,295 size 32x32
   Button "Button_61" at 39,328 size 32x32
   Button "Button_62" at 73,328 size 32x32
   Button "Button_63" at 107,328 size 32x32
   Button "Button_64" at 141,328 size 32x32
   Button "Button_65" at 175,328 size 32x32
   Button "Button_66" at 209,328 size 32x32
   Button "Button_67" at 243,328 size 32x32
   Button "Button_68" at 277,328 size 32x32
   Button "Button_69" at 311,328 size 32x32
   Button "Button_70" at 345,328 size 32x32
   Button "Button_71" at 39,361 size 32x32
   Button "Button_72" at 73,361 size 32x32
   Button "Button_73" at 107,361 size 32x32
   Button "Button_74" at 141,361 size 32x32
   Button "Button_75" at 175,361 size 32x32
   Button "Button_76" at 209,361 size 32x32
   Button "Button_77" at 243,361 size 32x32
   Button "Button_78" at 277,361 size 32x32
   Button "Button_79" at 311,361 size 32x32
   Button "Button_80" at 345,361 size 32x32
   Button "Button_81" at 39,394 size 32x32
   Button "Button_82" at 73,394 size 32x32
   Button "Button_83" at 107,394 size 32x32
   Button "Button_84" at 141,394 size 32x32
   Button "Button_85" at 175,394 size 32x32
   Button "Button_86" at 209,394 size 32x32
   Button "Button_87" at 243,394 size 32x32
   Button "Button_88" at 277,394 size 32x32
   Button "Button_89" at 311,394 size 32x32
   Button "Button_90" at 345,394 size 32x32
   Button "Button_91" at 39,427 size 32x32
   Button "Button_92" at 73,427 size 32x32
   Button "Button_93" at 107,427 size 32x32
   Button "Button_94" at 141,427 size 32x32
   Button "Button_95" at 175,427 size 32x32
   Button "Button_96" at 209,427 size 32x32
   Button "Button_97" at 243,427 size 32x32
   Button "Button_98" at 277,427 size 32x32
   Button "Button_99" at 311,427 size 32x32
   Button "Button_100" at 345,427 size 32x32
   GraphicView "Graphic view_2" at 410,97 size 376x366
   Button "Button_101" at 445,131 size 32x32
   Button "Button_102" at 479,131 size 32x32
   Button "Button_103" at 513,131 size 32x32
   Button "Button_104" at 547,131 size 32x32
   Button "Button_105" at 581,131 size 32x32
   Button "Button_106" at 615,131 size 32x32
   Button "Button_107" at 649,131 size 32x32
   Button "Button_108" at 683,131 size 32x32
   Button "Button_109" at 717,131 size 32x32
   Button "Button_110" at 751,131 size 32x32
   Button "Button_111" at 445,164 size 32x32
   Button "Button_112" at 479,164 size 32x32
   Button "Button_113" at 513,164 size 32x32
   Button "Button_114" at 547,164 size 32x32
   Button "Button_115" at 581,164 size 32x32
   Button "Button_116" at 615,164 size 32x32
   Button "Button_117" at 649,164 size 32x32
   Button "Button_118" at 683,164 size 32x32
   Button "Button_119" at 717,164 size 32x32
   Button "Button_120" at 751,164 size 32x32
   Button "Button_121" at 445,197 size 32x32
   Button "Button_122" at 479,197 size 32x32
   Button "Button_123" at 513,197 size 32x32
   Button "Button_124" at 547,197 size 32x32
   Button "Button_125" at 581,197 size 32x32
   Button "Button_126" at 615,197 size 32x32
   Button "Button_127" at 649,197 size 32x32
   Button "Button_128" at 683,197 size 32x32
   Button "Button_129" at 717,197 size 32x32
   Button "Button_130" at 751,197 size 32x32
   Button "Button_131" at 445,230 size 32x32
   Button "Button_132" at 479,230 size 32x32
   Button "Button_133" at 513,230 size 32x32
   Button "Button_134" at 547,230 size 32x32
   Button "Button_135" at 581,230 size 32x32
   Button "Button_136" at 615,230 size 32x32
   Button "Button_137" at 649,230 size 32x32
   Button "Button_138" at 683,230 size 32x32
   Button "Button_139" at 717,230 size 32x32
   Button "Button_140" at 751,230 size 32x32
   Button "Button_141" at 445,263 size 32x32
   Button "Button_142" at 479,263 size 32x32
   Button "Button_143" at 513,263 size 32x32
   Button "Button_144" at 547,263 size 32x32
   Button "Button_145" at 581,263 size 32x32
   Button "Button_146" at 615,263 size 32x32
   Button "Button_147" at 649,263 size 32x32
   Button "Button_148" at 683,263 size 32x32
   Button "Button_149" at 717,263 size 32x32
   Button "Button_150" at 751,263 size 32x32
   Button "Button_151" at 445,296 size 32x32
   Button "Button_152" at 479,296 size 32x32
   Button "Button_153" at 513,296 size 32x32
   Button "Button_154" at 547,296 size 32x32
   Button "Button_155" at 581,296 size 32x32
   Button "Button_156" at 615,296 size 32x32
   Button "Button_157" at 649,296 size 32x32
   Button "Button_158" at 683,296 size 32x32
   Button "Button_159" at 717,296 size 32x32
   Button "Button_160" at 751,296 size 32x32
   Button "Button_161" at 445,329 size 32x32
   Button "Button_162" at 479,329 size 32x32
   Button "Button_163" at 513,329 size 32x32
   Button "Button_164" at 547,329 size 32x32
   Button "Button_165" at 581,329 size 32x32
   Button "Button_166" at 615,329 size 32x32
   Button "Button_167" at 649,329 size 32x32
   Button "Button_168" at 683,329 size 32x32
   Button "Button_169" at 717,329 size 32x32
   Button "Button_170" at 751,329 size 32x32
   Button "Button_171" at 445,362 size 32x32
   Button "Button_172" at 479,362 size 32x32
   Button "Button_173" at 513,362 size 32x32
   Button "Button_174" at 547,362 size 32x32
   Button "Button_175" at 581,362 size 32x32
   Button "Button_176" at 615,362 size 32x32
   Button "Button_177" at 649,362 size 32x32
   Button "Button_178" at 683,362 size 32x32
   Button "Button_179" at 717,362 size 32x32
   Button "Button_180" at 751,362 size 32x32
   Button "Button_181" at 445,395 size 32x32
   Button "Button_182" at 479,395 size 32x32
   Button "Button_183" at 513,395 size 32x32
   Button "Button_184" at 547,395 size 32x32
   Button "Button_185" at 581,395 size 32x32
   Button "Button_186" at 615,395 size 32x32
   Button "Button_187" at 649,395 size 32x32
   Button "Button_188" at 683,395 size 32x32
   Button "Button_189" at 717,395 size 32x32
   Button "Button_190" at 751,395 size 32x32
   Button "Button_191" at 445,428 size 32x32
   Button "Button_192" at 479,428 size 32x32
   Button "Button_193" at 513,428 size 32x32
   Button "Button_194" at 547,428 size 32x32
   Button "Button_195" at 581,428 size 32x32
   Button "Button_196" at 615,428 size 32x32
   Button "Button_197" at 649,428 size 32x32
   Button "Button_198" at 683,428 size 32x32
   Button "Button_199" at 717,428 size 32x32
   Button "Button_200" at 751,428 size 32x32
*)